// TIA Portal project "ND_PiPl" (V16)
// Lehrlingsprojekt

(* hardware
DEVICE "ET 200SP-Station_1"  ET 200SP-Station
   slot 0: "Baugruppenträger_0"  Rack  6ES5 710-8MAx1
   slot 1: "-20KF3"  CPU 1512SP F-1 PN  6ES7 512-1SK01-0AB0  V2.8
      slot 32768: "PROFINET-Schnittstelle_1"  X1
         slot 32771: "Port_3"  X1 P3
   slot 2: "-20KF5"  F-DI 8x24VDC HF  6ES7 136-6BA00-0CA0  V1.0
      slot 1: "-20KF5"  F-DI 8x24VDC HF
   slot 3: "-20KF6"  F-DQ 8x24VDC/0.5A PP HF  6ES7 136-6DC00-0CA0  V1.0
      slot 1: "-20KF6"  F-DQ 8x24VDC/0.5A PP HF
   slot 4: "-21KF1"  DI 16x24VDC ST  6ES7 131-6BH01-0BA0  V0.0
      slot 1: "-21KF1"  DI 16x24VDC ST
   slot 5: "-21KF4"  DQ 16x24VDC/0.5A ST  6ES7 132-6BH01-0BA0  V0.0
      slot 1: "-21KF4"  DQ 16x24VDC/0.5A ST
   slot 6: "-22KF1"  AI 2xU/I 2-,4-wire HS  6ES7 134-6HB00-0DA1  V2.0
      slot 1: "-22KF1"  AI 2xU/I 2-,4-wire HS
   slot 7: "-22KF3"  AQ 2xU ST  6ES7 135-6FB00-0BA1  V1.0
      slot 1: "-22KF3"  AQ 2xU ST
   slot 8: "Servermodul_1"  Server module  6ES7 193-6PA00-0AA0  V1.1
      slot 1: "Servermodul_1"  Server module
   slot 127: "BA 2xRJ45"  BA 2xRJ45  6ES7 193-6AR00-0AA0  V0.0
      slot 32769: "Port_1"  X1 P1  6ES7 193-6AR00-0AA0
      slot 32770: "Port_2"  X1 P2  6ES7 193-6AR00-0AA0
DEVICE "HMI_1"  KTP400 Comfort
   slot 0: "HMI_1"  KTP400 Comfort  6AV2 124-2DC01-0AX0  16.0.0.0
   slot 1: "HMI_RT_1"  KTP400 Comfort  6AV2 124-2DC01-0AX0  16.0.0.0
   slot 5: "HMI_1.IE_CP_1"  PROFINET Interface  16.0.0.0
      slot 1: "PROFINET Schnittstelle_1"  PROFINET Interface
         slot 1: "Port_1"  Port
   slot 7: "HMI_1.MPI/DP_CP_1"  MPI/DP Interface  16.0.0.0
*)

// ===== PLC "-20KF3"  CPU 1512SP F-1 PN =====
// protected blocks, not shown: "Main_Safety_RTG1", "Main_Safety_RTG1_DB"

VAR_GLOBAL   // PLC tag table "Standard-Variablentabelle"
   "FirstScan" AT %M1.0 : Bool;
   "DiagStatusUpdate" AT %M1.1 : Bool;
   "AlwaysTRUE" AT %M1.2 : Bool;
   "AlwaysFALSE" AT %M1.3 : Bool;
   "Clock_10Hz" AT %M50.0 : Bool;
   "Clock_5Hz" AT %M50.1 : Bool;
   "Clock_2.5Hz" AT %M50.2 : Bool;
   "Clock_2Hz" AT %M50.3 : Bool;
   "Clock_1.25Hz" AT %M50.4 : Bool;
   "Clock_1Hz" AT %M50.5 : Bool;
   "Clock_0.625Hz" AT %M50.6 : Bool;
   "Clock_0.5Hz" AT %M50.7 : Bool;
   "MaschineStart" AT %M900.0 : Bool;
   "Schritt_Förderband_Ein" AT %M900.1 : Bool;
   "Schritt_Vereinzelner_Ein" AT %M900.2 : Bool;
   "Vereinzler_Ein" AT %M1000.0 : Bool;
   "Schritt_Horizontalarm_Zurück" AT %M900.3 : Bool;
   "Schritt_Vakuum_Ein" AT %M900.4 : Bool;
   "VakuumSR" AT %M1000.1 : Bool;
   "Förderband_Merker" AT %M2000.0 : Bool;
   "Schritt_Vertikalarm_runter" AT %M900.5 : Bool;
   "Tag_2" AT %M1000.2 : Bool;
   "Schritt_Vertikalarm_oben" AT %M900.6 : Bool;
   "Schritt_Horizontalarm_vor" AT %M900.7 : Bool;
   "Schritt_VertikalarmDeckel_runter" AT %M901.0 : Bool;
   "Schritt_Vakuum_aus" AT %M901.1 : Bool;
   "Schritt_VertikalarmDeckelweg_oben" AT %M901.2 : Bool;
   "Schritt_HorizontalarmDeckel_zurück" AT %M901.3 : Bool;
   "Schritt_Vereinzler_aus" AT %M901.4 : Bool;
   "Schritt_Zurücksetzten_Anfang" AT %M901.5 : Bool;
   "Start_Impuls" AT %M200.1 : Bool;
   "Einmal_Start" AT %M2000.1 : Bool;
   "Stop_Speicher" AT %M2000.2 : Bool;
   "Deckler_Speicher" AT %M2000.3 : Bool;
   "Tag_1" AT %ED500 : Real;
   "Druck_Zu_Niedrig" AT %M2000.4 : Bool;
   "Druck_Zu_Hoch" AT %M2000.5 : Bool;
   "Prod_Count" AT %MW1200 : Int;
   "Prod_Count_Reset" AT %M300.0 : Bool;
END_VAR

VAR_GLOBAL   // PLC tag table "Systemflags"
   "System_Byte" AT %MB1 : Byte;   // Byte System
   "ME_PLC_First_Scan_Bit" AT %M1.0 : Bool;   // PLC First Scan Bit
   "ME_PLC_DiagStatusUpdate" AT %M1.1 : Bool;   // PLC Diagnostic Status Update
   "ME_PLC_TRUE" AT %M1.2 : Bool;   // PLC TRUE
   "ME_PLC_FALSE" AT %M1.3 : Bool;   // PLC FALSE
   "Clock_Byte" AT %MB50 : Byte;   // Byte PLC Clock
   "ME_PLC_Clock_0.1s" AT %M0.0 : Bool;   // PLC Clock 0.1s (10Hz )
   "ME_PLC_Clock_0.2s" AT %M0.1 : Bool;   // PLC Clock 0.2s (5Hz )
   "ME_PLC_Clock_0.4s" AT %M0.2 : Bool;   // PLC Clock 0.4s (2.5Hz )
   "ME_PLC_Clock_0.5s" AT %M0.3 : Bool;   // PLC Clock 0.5s (2Hz )
   "ME_PLC_Clock_0.8s" AT %M0.4 : Bool;   // PLC Clock 0.8s (1.25Hz )
   "ME_PLC_Clock_1.0s" AT %M0.5 : Bool;   // PLC Clock 1s (1Hz)
   "ME_PLC_Clock_1.6s" AT %M0.6 : Bool;   // PLC Clock 1.6s (0.625Hz )
   "ME_PLC_Clock_2.0s" AT %M0.7 : Bool;   // PLC Clock 2s (0.5Hz )
   "ME_PLC_FC_Test" AT %M2.0 : Bool;   // Testing Frequency Converters
   "ME_PLC_TRUE_to_do" AT %M2.2 : Bool;   // PLC TRUE to do
   "ME_PLC_FALSE_to_do" AT %M2.3 : Bool;   // PLC FALSE to do
   "ME_PLC_Led_Error" AT %M2.4 : Bool;   // PLC LED Error
   "ME_PLC_Led_Maint" AT %M2.5 : Bool;   // PLC LED Maintenance
   "ME_PLC_Startup_Rst" AT %M2.6 : Bool;   // PLC LED Startup Reset
   "ME_PLC_First_Scan_Bit_FC" AT %M2.1 : Bool;   // Call Frequency Converters
END_VAR

VAR_GLOBAL   // PLC tag table "IO-Pick&Placer"
   "CC_KF_FbEStop" AT %E0.0 : Bool;   // Rückmeldung Freigabe Not-Halt (81KF8)
   "PPTR_BG_InletPart" AT %E0.1 : Bool;   // Transportband Werkstück am Bandanfang (100BG1)
   "PPTR_BG_PartAtSep" AT %E0.2 : Bool;   // Transportband Werkstück am Vereinzeler (100BG2)
   "PPTR_BG_BackupPart" AT %E0.3 : Bool;   // Transportband Werkstück beim Bandende (100BG3)
   "PIPL_BG_CarrierRetracted" AT %E0.4 : Bool;   // Pick&Placer Schlitten eingefahren (120BG1)
   "PIPL_BG_CarrierExtended" AT %E0.5 : Bool;   // Pick&Placer Schlitten ausgefahren (120BG2)
   "PIPL_BG_SuctTop" AT %E0.6 : Bool;   // Pick&Placer Sauger oben (120BG3)
   "PIPL_BP_PartSuckedOn" AT %E0.7 : Bool;   // Pick&Placer Werkstück angesaugt (120PB4)
   "PIPL_Pa_SF_Reset" AT %E1.0 : Bool;   // Pick&Placer Bedienstelle Reset (160SF2)
   "PIPL_Pa_SF_Start" AT %E1.1 : Bool;   // Pick&Placer Bedienstelle Start (160SF3)
   "PIPL_Pa_SF_Stop" AT %E1.2 : Bool;   // Pick&Placer Bedienstelle Stop (160SF4)
   "PIPL_Pa_SF_ManAuto" AT %E1.3 : Bool;   // Pick&Placer Bedienstelle Manual - Auto (160SF5)
   "CC_Spare_I1.4" AT %E1.4 : Bool;   // Spare
   "CC_Spare_I1.5" AT %E1.5 : Bool;   // Spare
   "CC_Spare_I1.6" AT %E1.6 : Bool;   // Spare
   "CC_Spare_I1.7" AT %E1.7 : Bool;   // Spare
   "PPTR_MB_SeparatorExtend" AT %A0.0 : Bool;   // Transportband Vereinzeler ausfahren (105MB8)
   "PIPL_SC_Green" AT %A0.1 : Bool;   // Pick&Placer Turmleuchte grün (130PF1)
   "PIPL_SC_Yellow" AT %A0.2 : Bool;   // Pick&Placer Turmleuchte gelb (130PF1)
   "PIPL_SC_Red" AT %A0.3 : Bool;   // Pick&Placer Turmleuchte rot (130PF1)
   "PIPL_MB_CarrierExtend" AT %A0.4 : Bool;   // Pick&Placer Schlitten ausfahren (125MB1)
   "PIPL_MB_CarrierRetract" AT %A0.5 : Bool;   // Pick&Placer Schlitten einfahren (125MB2)
   "PIPL_MB_SuctDown" AT %A0.6 : Bool;   // Pick&Placer Sauger nach unten (125MB3)
   "PIPL_MB_VacuumOn" AT %A0.7 : Bool;   // Pick&Placer Vakuum ein (125MB4)
   "PIPL_Pa_PF_ControlCircuit" AT %A1.0 : Bool;   // Pick&Placer Bedienstelle LED Steuerspannung Ein (Reset) (160SF2)
   "PIPL_Pa_PF_Error" AT %A1.1 : Bool;   // Pick&Placer Bedienstelle LED Fehler (160PF2)
   "PIPL_Pa_PF_Start" AT %A1.2 : Bool;   // Pick&Placer Bedienstelle LED Start (160SF3)
   "CC_Spare_O1.3" AT %A1.3 : Bool;   // Spare
   "CC_Spare_O1.4" AT %A1.4 : Bool;   // Spare
   "CC_Spare_O1.5" AT %A1.5 : Bool;   // Spare
   "CC_Spare_O1.6" AT %A1.6 : Bool;   // Spare
   "CC_Spare_O1.7" AT %A1.7 : Bool;   // Spare
   "Druck_Tester" AT %EW272 : Int;   // Druck Tester
   "CC_Spare_IW274" AT %EW274 : Word;   // Spare
   "PPTR_TF_DriveSpeed" AT %AW272 : Word;   // Transportband Bandmotor Geschwindigkeit Option (105TF1)
   "CC_Spare_OW274" AT %AW274 : Word;   // Spare
   "Druck_Zwischenwert" AT %MD276 : Real;
   "Druck_Wert1" AT %MD280 : Real;
   "Druck_Wert2" AT %MW284 : Int;
   "Druck_Wert_Final" AT %MD286 : Real;
END_VAR

VAR_GLOBAL   // PLC tag table "IO-Pick&Placer-Safety"
   "PIPL_Pa_EStopCh1" AT %E1000.0 : Bool;   // Pick&Placer Bedienstelle Not-Halt Channel 1 (160SF1)
   "CC_Spare_I1000.1" AT %E1000.1 : Bool;   // Spare
   "CC_Spare_I1000.2" AT %E1000.2 : Bool;   // Spare
   "CC_Spare_I1000.3" AT %E1000.3 : Bool;   // Spare
   "PIPL_Pa_EStopCh2" AT %E1000.4 : Bool;   // Pick&Placer Bedienstelle Not-Halt Channel 2 (160SF1)
   "CC_Spare_I1000.5" AT %E1000.5 : Bool;   // Spare
   "CC_Spare_I1000.6" AT %E1000.6 : Bool;   // Spare
   "CC_Spare_I1000.7" AT %E1000.7 : Bool;   // Spare
   "CC_KF_EStopCh1" AT %A1050.0 : Bool;   // Freigabe Not-Halt Channel 1 (81KF7)
   "CC_KF_EStopCh2" AT %A1050.1 : Bool;   // Freigabe Not-Halt Channel 2 (81KF8)
   "PPTR_TF_DriveForward" AT %A1050.2 : Bool;   // Transportband Bandmotor Vorwärts (105TF1)
   "PPTR_TF_DriveReverse" AT %A1050.3 : Bool;   // Transportband Bandmotor Rückwärts (105TF1)
   "CC_Spare_O1050.4" AT %A1050.4 : Bool;   // Spare
   "CC_Spare_O1050.5" AT %A1050.5 : Bool;   // Spare
   "CC_Spare_O1050.6" AT %A1050.6 : Bool;   // Spare
   "CC_Spare_O1050.7" AT %A1050.7 : Bool;   // Spare
END_VAR

DATA_BLOCK "HMI_Meldungen"   // DB120
{ S7_Optimized_Access := 'FALSE' }
VERSION : 0.1
   VAR
      Fehler : Struct
         "Not-Aus" : Bool;   // NOT-Aus Aktiv
         "Not-Aus_Quit" : Bool;   // NOT-Aus Quitieren
         "2" : Bool;
         "3" : Bool;
         "4" : Bool;
         "5" : Bool;
         "6" : Bool;
         "7" : Bool;
         "8" : Bool;
         "9" : Bool;
         "10" : Bool;
         "11" : Bool;
         "12" : Bool;
         "13" : Bool;
         "14" : Bool;
         "15" : Bool;
      END_STRUCT;
      Meldungen : Struct
         "0" : Bool;
         "1" : Bool;
         "2" : Bool;
         "3" : Bool;
         "4" : Bool;
         "5" : Bool;
         "6" : Bool;
         "7" : Bool;
         "8" : Bool;
         "9" : Bool;
         "10" : Bool;
         "11" : Bool;
         "12" : Bool;
         "13" : Bool;
         "14" : Bool;
         "15" : Bool;
      END_STRUCT;
      Warnungen : Struct
         Druck_zu_niedrig : Bool;   // Druck zu niedrig
         Druck_zu_hoch : Bool;   // Druck zu hoch
         Keine_Deckel : Bool;   // Keine Deckel vorhanden
         Rückstau : Bool;   // Rückstau am Bandende
         "4" : Bool;
         "5" : Bool;
         "6" : Bool;
         "7" : Bool;
         "8" : Bool;
         "9" : Bool;
         "10" : Bool;
         "11" : Bool;
         "12" : Bool;
         "13" : Bool;
         "14" : Bool;
         "15" : Bool;
      END_STRUCT;
   END_VAR
BEGIN
END_DATA_BLOCK

// folder: System blocks/Program resources

DATA_BLOCK "IEC_Timer_0_DB"   // DB3
{ S7_Optimized_Access := 'TRUE' }
AUTHOR : Simatic
FAMILY : IEC
NAME : IEC_TMR
VERSION : 1.0
// stored: InstanceOfName IEC_TIMER
"IEC_TIMER"
BEGIN
END_DATA_BLOCK

DATA_BLOCK "Vakuum_Timer_Ausschalten"   // DB5
{ S7_Optimized_Access := 'TRUE' }
AUTHOR : Simatic
FAMILY : IEC
NAME : IEC_TMR
VERSION : 1.0
// stored: InstanceOfName IEC_TIMER
"IEC_TIMER"
BEGIN
END_DATA_BLOCK

DATA_BLOCK "Timer_Rückstau"   // DB6
{ S7_Optimized_Access := 'TRUE' }
AUTHOR : Simatic
FAMILY : IEC
NAME : IEC_TMR
VERSION : 1.0
// stored: InstanceOfName IEC_TIMER
"IEC_TIMER"
BEGIN
END_DATA_BLOCK

DATA_BLOCK "Timer_Clean_Reset"   // DB7
{ S7_Optimized_Access := 'TRUE' }
AUTHOR : Simatic
FAMILY : IEC
NAME : IEC_TMR
VERSION : 1.0
// stored: InstanceOfName IEC_TIMER
"IEC_TIMER"
BEGIN
END_DATA_BLOCK

DATA_BLOCK "IEC_Counter_0_DB"   // DB8
{ S7_Optimized_Access := 'TRUE' }
AUTHOR : Simatic
FAMILY : IEC
NAME : CNTR
VERSION : 1.0
// stored: InstanceOfName IEC_COUNTER
"IEC_COUNTER"
BEGIN
END_DATA_BLOCK

// folder: (top level)

FUNCTION "Ausgänge" : Void   // FC1, FBD
{ S7_Optimized_Access := 'TRUE' }
VERSION : 0.1
BEGIN

REGION Network 1: Vereinzler
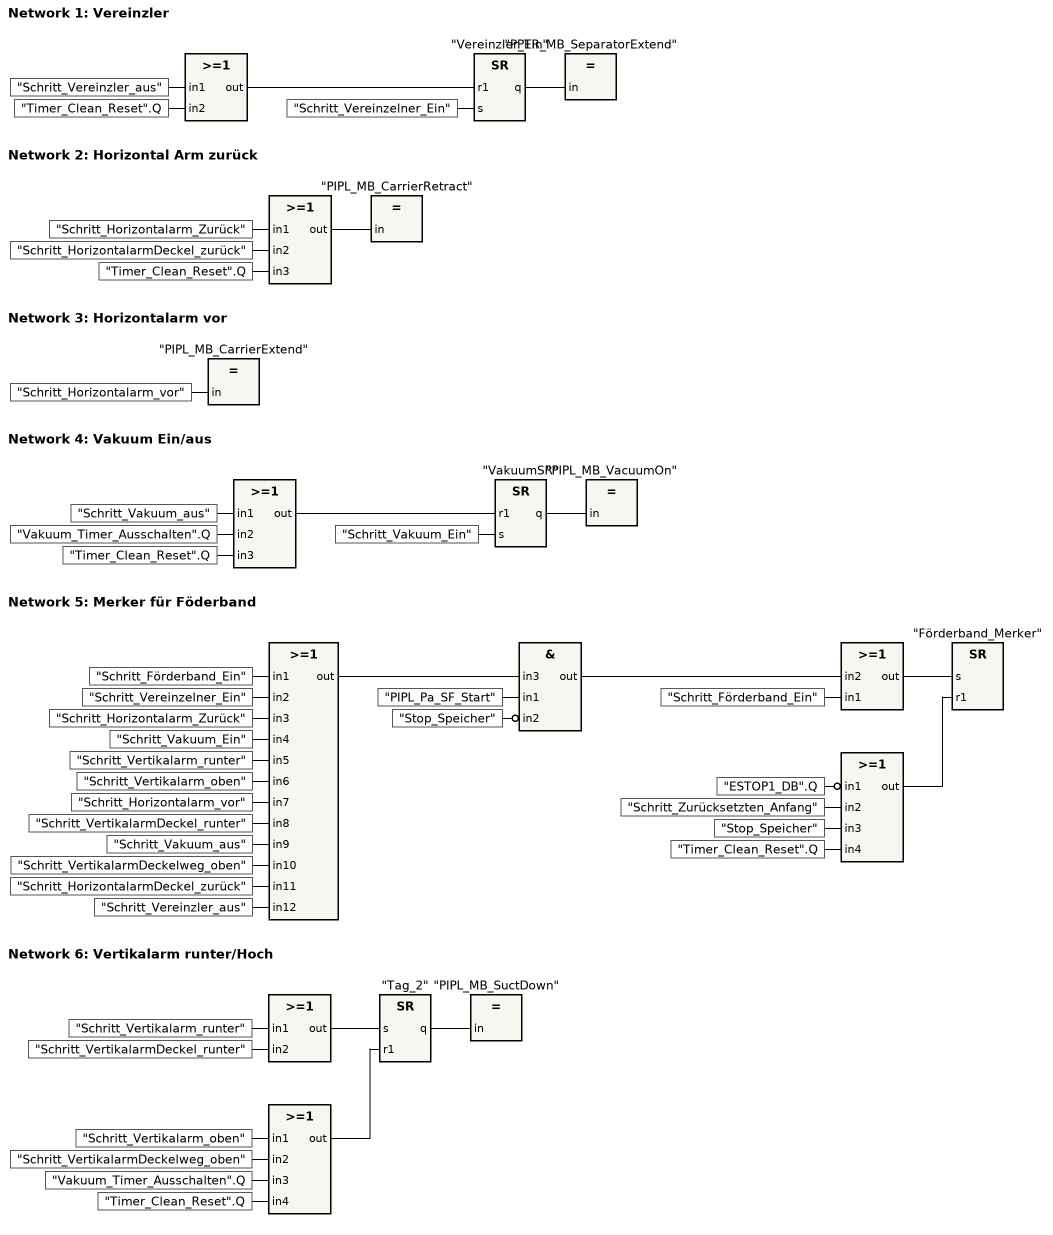
   IF "Schritt_Vereinzelner_Ein" THEN
       "Vereinzler_Ein" := TRUE;   // SR flip-flop
   END_IF;
   IF "Schritt_Vereinzler_aus" OR "Timer_Clean_Reset".Q THEN "Vereinzler_Ein" := FALSE; END_IF;
   "PPTR_MB_SeparatorExtend" := "Vereinzler_Ein";
END_REGION

REGION Network 2: Horizontal Arm zurück
   "PIPL_MB_CarrierRetract" := "Schritt_Horizontalarm_Zurück" OR "Schritt_HorizontalarmDeckel_zurück" OR "Timer_Clean_Reset".Q;
END_REGION

REGION Network 3: Horizontalarm vor
   "PIPL_MB_CarrierExtend" := "Schritt_Horizontalarm_vor";
END_REGION

REGION Network 4: Vakuum Ein/aus
   IF "Schritt_Vakuum_Ein" THEN
       "VakuumSR" := TRUE;   // SR flip-flop
   END_IF;
   IF "Schritt_Vakuum_aus" OR "Vakuum_Timer_Ausschalten".Q OR "Timer_Clean_Reset".Q THEN
       "VakuumSR" := FALSE;
   END_IF;
   "PIPL_MB_VacuumOn" := "VakuumSR";
END_REGION

REGION Network 5: Merker für Föderband
   IF (("Schritt_Förderband_Ein" OR "Schritt_Vereinzelner_Ein" OR "Schritt_Horizontalarm_Zurück" OR "Schritt_Vakuum_Ein" OR "Schritt_Vertikalarm_runter" OR "Schritt_Vertikalarm_oben" OR "Schritt_Horizontalarm_vor" OR "Schritt_VertikalarmDeckel_runter" OR "Schritt_Vakuum_aus" OR "Schritt_VertikalarmDeckelweg_oben" OR "Schritt_HorizontalarmDeckel_zurück" OR "Schritt_Vereinzler_aus") AND "PIPL_Pa_SF_Start" AND NOT "Stop_Speicher") OR "Schritt_Förderband_Ein" THEN
       "Förderband_Merker" := TRUE;   // SR flip-flop
   END_IF;
   IF NOT "ESTOP1_DB".Q OR "Schritt_Zurücksetzten_Anfang" OR "Stop_Speicher" OR "Timer_Clean_Reset".Q THEN
       "Förderband_Merker" := FALSE;
   END_IF;
END_REGION

REGION Network 6: Vertikalarm runter/Hoch
   IF "Schritt_Vertikalarm_runter" OR "Schritt_VertikalarmDeckel_runter" THEN
       "Tag_2" := TRUE;   // SR flip-flop
   END_IF;
   IF "Schritt_Vertikalarm_oben" OR "Schritt_VertikalarmDeckelweg_oben" OR "Vakuum_Timer_Ausschalten".Q OR "Timer_Clean_Reset".Q THEN
       "Tag_2" := FALSE;
   END_IF;
   "PIPL_MB_SuctDown" := "Tag_2";
END_REGION
END_FUNCTION

FUNCTION "Pick&Place_Auto" : Void   // FC2, FBD
{ S7_Optimized_Access := 'TRUE' }
VERSION : 0.1
BEGIN

REGION Network 1: Eischalten der Maschine
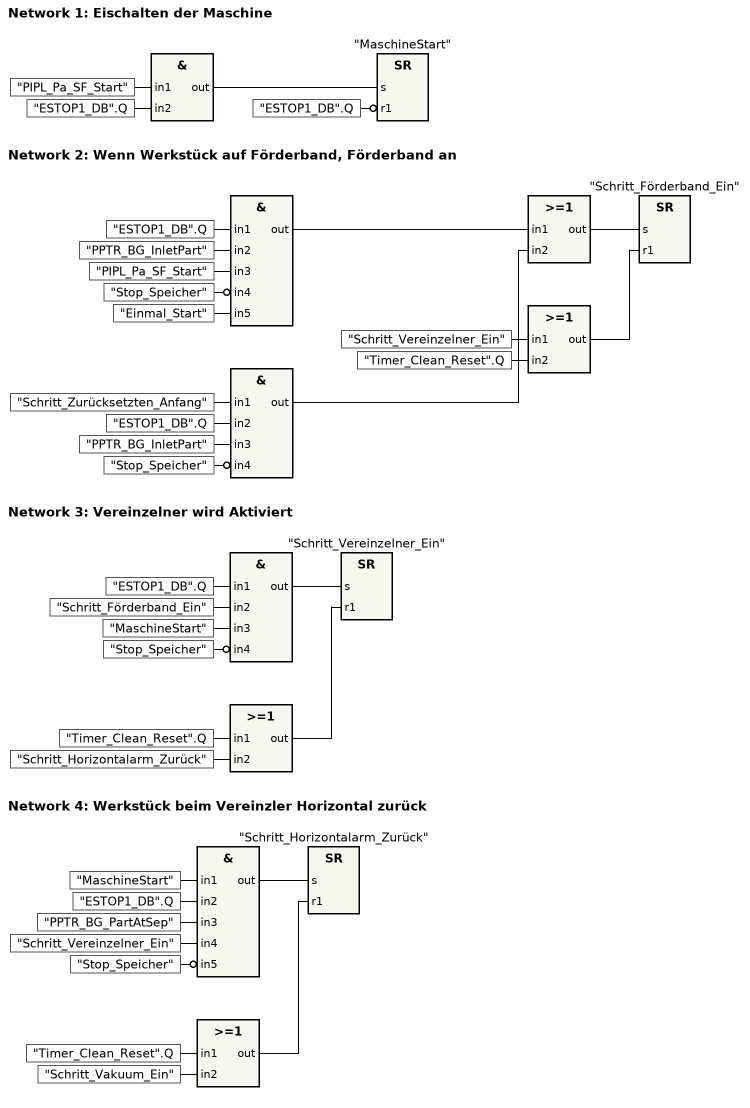
   IF "PIPL_Pa_SF_Start" AND "ESTOP1_DB".Q THEN
       "MaschineStart" := TRUE;   // SR flip-flop
   END_IF;
   IF NOT "ESTOP1_DB".Q THEN "MaschineStart" := FALSE; END_IF;
END_REGION

REGION Network 2: Wenn Werkstück auf Förderband, Förderband an
   IF ("ESTOP1_DB".Q AND "PPTR_BG_InletPart" AND "PIPL_Pa_SF_Start" AND NOT "Stop_Speicher" AND "Einmal_Start") OR ("Schritt_Zurücksetzten_Anfang" AND "ESTOP1_DB".Q AND "PPTR_BG_InletPart" AND NOT "Stop_Speicher") THEN
       "Schritt_Förderband_Ein" := TRUE;   // SR flip-flop
   END_IF;
   IF "Schritt_Vereinzelner_Ein" OR "Timer_Clean_Reset".Q THEN "Schritt_Förderband_Ein" := FALSE; END_IF;
END_REGION

REGION Network 3: Vereinzelner wird Aktiviert
   IF "ESTOP1_DB".Q AND "Schritt_Förderband_Ein" AND "MaschineStart" AND NOT "Stop_Speicher" THEN
       "Schritt_Vereinzelner_Ein" := TRUE;   // SR flip-flop
   END_IF;
   IF "Timer_Clean_Reset".Q OR "Schritt_Horizontalarm_Zurück" THEN
       "Schritt_Vereinzelner_Ein" := FALSE;
   END_IF;
END_REGION

REGION Network 4: Werkstück beim Vereinzler Horizontal zurück
   IF "MaschineStart" AND "ESTOP1_DB".Q AND "PPTR_BG_PartAtSep" AND "Schritt_Vereinzelner_Ein" AND NOT "Stop_Speicher" THEN
       "Schritt_Horizontalarm_Zurück" := TRUE;   // SR flip-flop
   END_IF;
   IF "Timer_Clean_Reset".Q OR "Schritt_Vakuum_Ein" THEN "Schritt_Horizontalarm_Zurück" := FALSE; END_IF;
END_REGION

REGION Network 5: Wenn Horizontalarm zurück, Vakuum ein
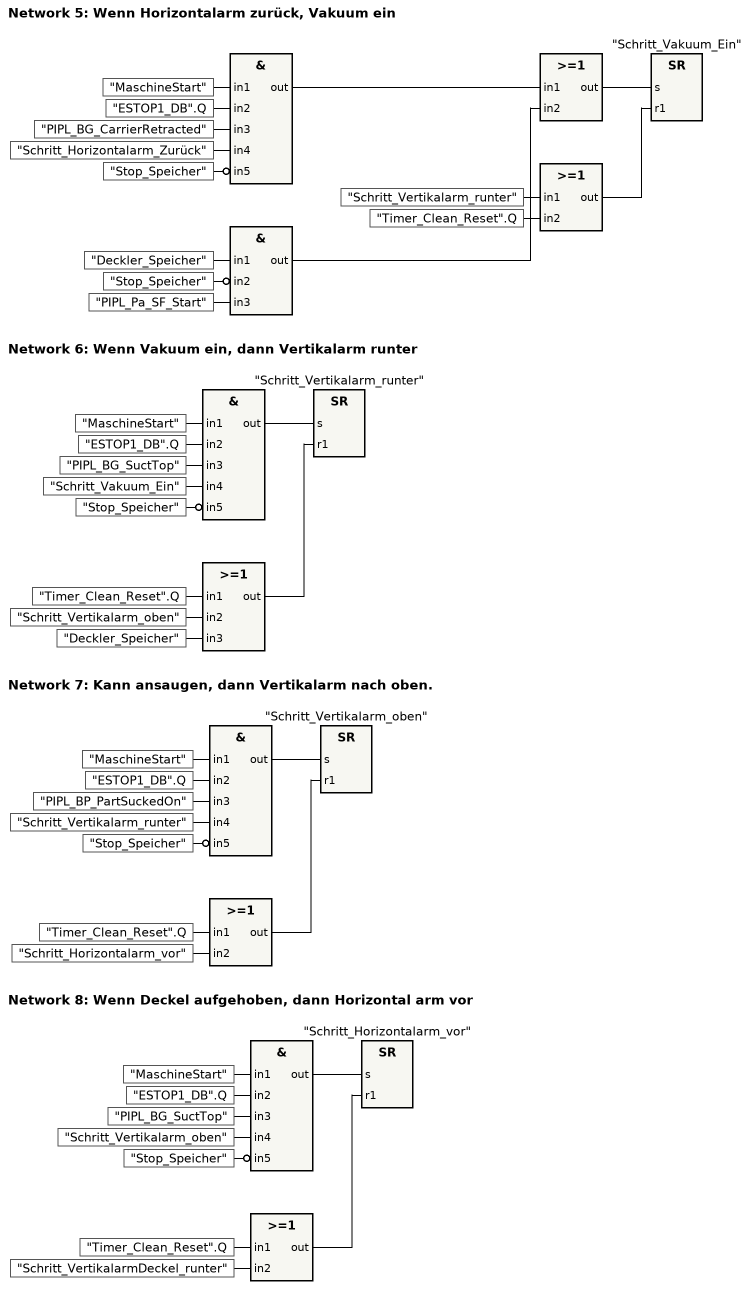
   IF ("MaschineStart" AND "ESTOP1_DB".Q AND "PIPL_BG_CarrierRetracted" AND "Schritt_Horizontalarm_Zurück" AND NOT "Stop_Speicher") OR ("Deckler_Speicher" AND NOT "Stop_Speicher" AND "PIPL_Pa_SF_Start") THEN
       "Schritt_Vakuum_Ein" := TRUE;   // SR flip-flop
   END_IF;
   IF "Schritt_Vertikalarm_runter" OR "Timer_Clean_Reset".Q THEN "Schritt_Vakuum_Ein" := FALSE; END_IF;
END_REGION

REGION Network 6: Wenn Vakuum ein, dann Vertikalarm runter
   IF "MaschineStart" AND "ESTOP1_DB".Q AND "PIPL_BG_SuctTop" AND "Schritt_Vakuum_Ein" AND NOT "Stop_Speicher" THEN
       "Schritt_Vertikalarm_runter" := TRUE;   // SR flip-flop
   END_IF;
   IF "Timer_Clean_Reset".Q OR "Schritt_Vertikalarm_oben" OR "Deckler_Speicher" THEN
       "Schritt_Vertikalarm_runter" := FALSE;
   END_IF;
END_REGION

REGION Network 7: Kann ansaugen, dann Vertikalarm nach oben.
   IF "MaschineStart" AND "ESTOP1_DB".Q AND "PIPL_BP_PartSuckedOn" AND "Schritt_Vertikalarm_runter" AND NOT "Stop_Speicher" THEN
       "Schritt_Vertikalarm_oben" := TRUE;   // SR flip-flop
   END_IF;
   IF "Timer_Clean_Reset".Q OR "Schritt_Horizontalarm_vor" THEN "Schritt_Vertikalarm_oben" := FALSE; END_IF;
END_REGION

REGION Network 8: Wenn Deckel aufgehoben, dann Horizontal arm vor
   IF "MaschineStart" AND "ESTOP1_DB".Q AND "PIPL_BG_SuctTop" AND "Schritt_Vertikalarm_oben" AND NOT "Stop_Speicher" THEN
       "Schritt_Horizontalarm_vor" := TRUE;   // SR flip-flop
   END_IF;
   IF "Timer_Clean_Reset".Q OR "Schritt_VertikalarmDeckel_runter" THEN
       "Schritt_Horizontalarm_vor" := FALSE;
   END_IF;
END_REGION

REGION Network 9: Wenn Horizontalarm vor mit Deckel, dann Vertickalarm runter
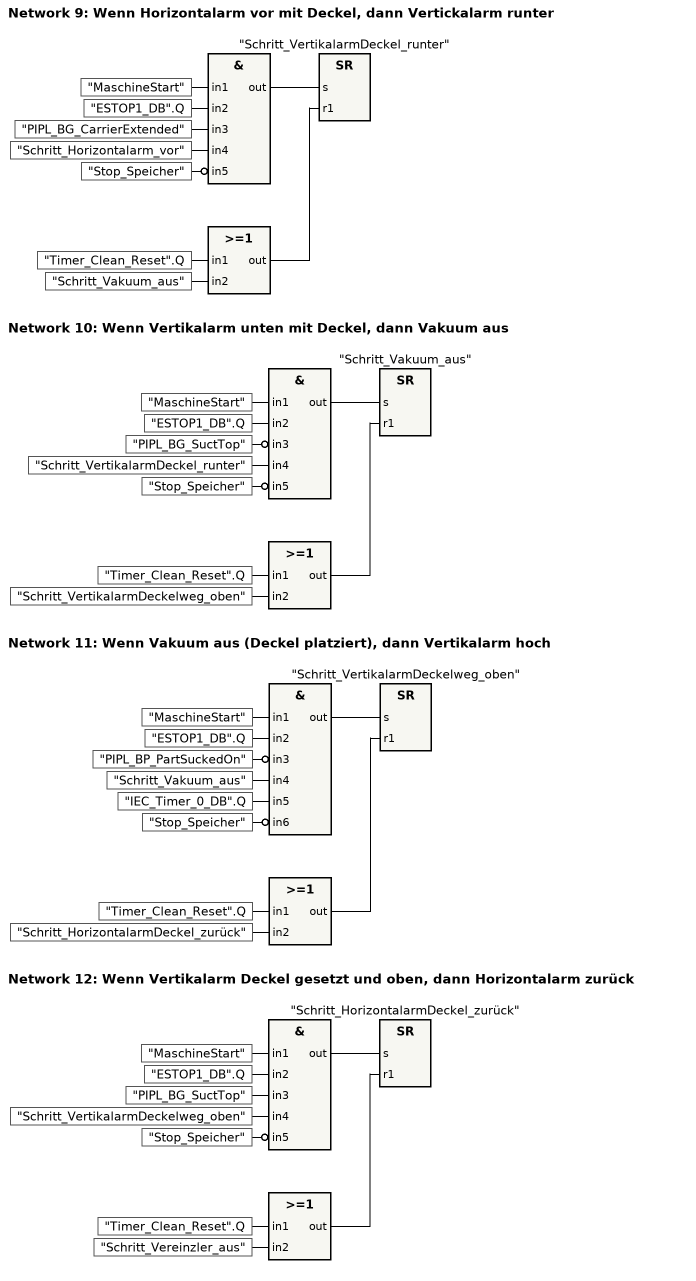
   IF "MaschineStart" AND "ESTOP1_DB".Q AND "PIPL_BG_CarrierExtended" AND "Schritt_Horizontalarm_vor" AND NOT "Stop_Speicher" THEN
       "Schritt_VertikalarmDeckel_runter" := TRUE;   // SR flip-flop
   END_IF;
   IF "Timer_Clean_Reset".Q OR "Schritt_Vakuum_aus" THEN "Schritt_VertikalarmDeckel_runter" := FALSE; END_IF;
END_REGION

REGION Network 10: Wenn Vertikalarm unten mit Deckel, dann Vakuum aus
   IF "MaschineStart" AND "ESTOP1_DB".Q AND NOT "PIPL_BG_SuctTop" AND "Schritt_VertikalarmDeckel_runter" AND NOT "Stop_Speicher" THEN
       "Schritt_Vakuum_aus" := TRUE;   // SR flip-flop
   END_IF;
   IF "Timer_Clean_Reset".Q OR "Schritt_VertikalarmDeckelweg_oben" THEN
       "Schritt_Vakuum_aus" := FALSE;
   END_IF;
END_REGION

REGION Network 11: Wenn Vakuum aus (Deckel platziert), dann Vertikalarm hoch
   IF "MaschineStart" AND "ESTOP1_DB".Q AND NOT "PIPL_BP_PartSuckedOn" AND "Schritt_Vakuum_aus" AND "IEC_Timer_0_DB".Q AND NOT "Stop_Speicher" THEN
       "Schritt_VertikalarmDeckelweg_oben" := TRUE;   // SR flip-flop
   END_IF;
   IF "Timer_Clean_Reset".Q OR "Schritt_HorizontalarmDeckel_zurück" THEN
       "Schritt_VertikalarmDeckelweg_oben" := FALSE;
   END_IF;
END_REGION

REGION Network 12: Wenn Vertikalarm Deckel gesetzt und oben, dann Horizontalarm zurück
   IF "MaschineStart" AND "ESTOP1_DB".Q AND "PIPL_BG_SuctTop" AND "Schritt_VertikalarmDeckelweg_oben" AND NOT "Stop_Speicher" THEN
       "Schritt_HorizontalarmDeckel_zurück" := TRUE;   // SR flip-flop
   END_IF;
   IF "Timer_Clean_Reset".Q OR "Schritt_Vereinzler_aus" THEN
       "Schritt_HorizontalarmDeckel_zurück" := FALSE;
   END_IF;
END_REGION

REGION Network 13: Wenn Horizontalarm zurück (Deckel platziert), dann Vereinzler aus
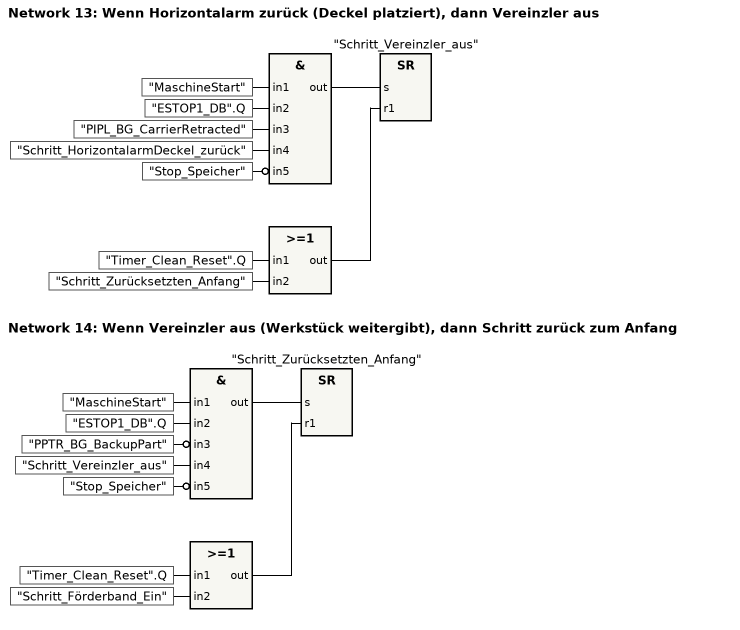
   IF "MaschineStart" AND "ESTOP1_DB".Q AND "PIPL_BG_CarrierRetracted" AND "Schritt_HorizontalarmDeckel_zurück" AND NOT "Stop_Speicher" THEN
       "Schritt_Vereinzler_aus" := TRUE;   // SR flip-flop
   END_IF;
   IF "Timer_Clean_Reset".Q OR "Schritt_Zurücksetzten_Anfang" THEN "Schritt_Vereinzler_aus" := FALSE; END_IF;
END_REGION

REGION Network 14: Wenn Vereinzler aus (Werkstück weitergibt), dann Schritt zurück zum Anfang
   IF "MaschineStart" AND "ESTOP1_DB".Q AND NOT "PPTR_BG_BackupPart" AND "Schritt_Vereinzler_aus" AND NOT "Stop_Speicher" THEN
       "Schritt_Zurücksetzten_Anfang" := TRUE;   // SR flip-flop
   END_IF;
   IF "Timer_Clean_Reset".Q OR "Schritt_Förderband_Ein" THEN "Schritt_Zurücksetzten_Anfang" := FALSE; END_IF;
END_REGION
END_FUNCTION

FUNCTION "SonderBlöcke" : Void   // FC3, FBD
{ S7_Optimized_Access := 'TRUE' }
VERSION : 0.1
BEGIN

REGION Network 1: Delay für Deckel setzen
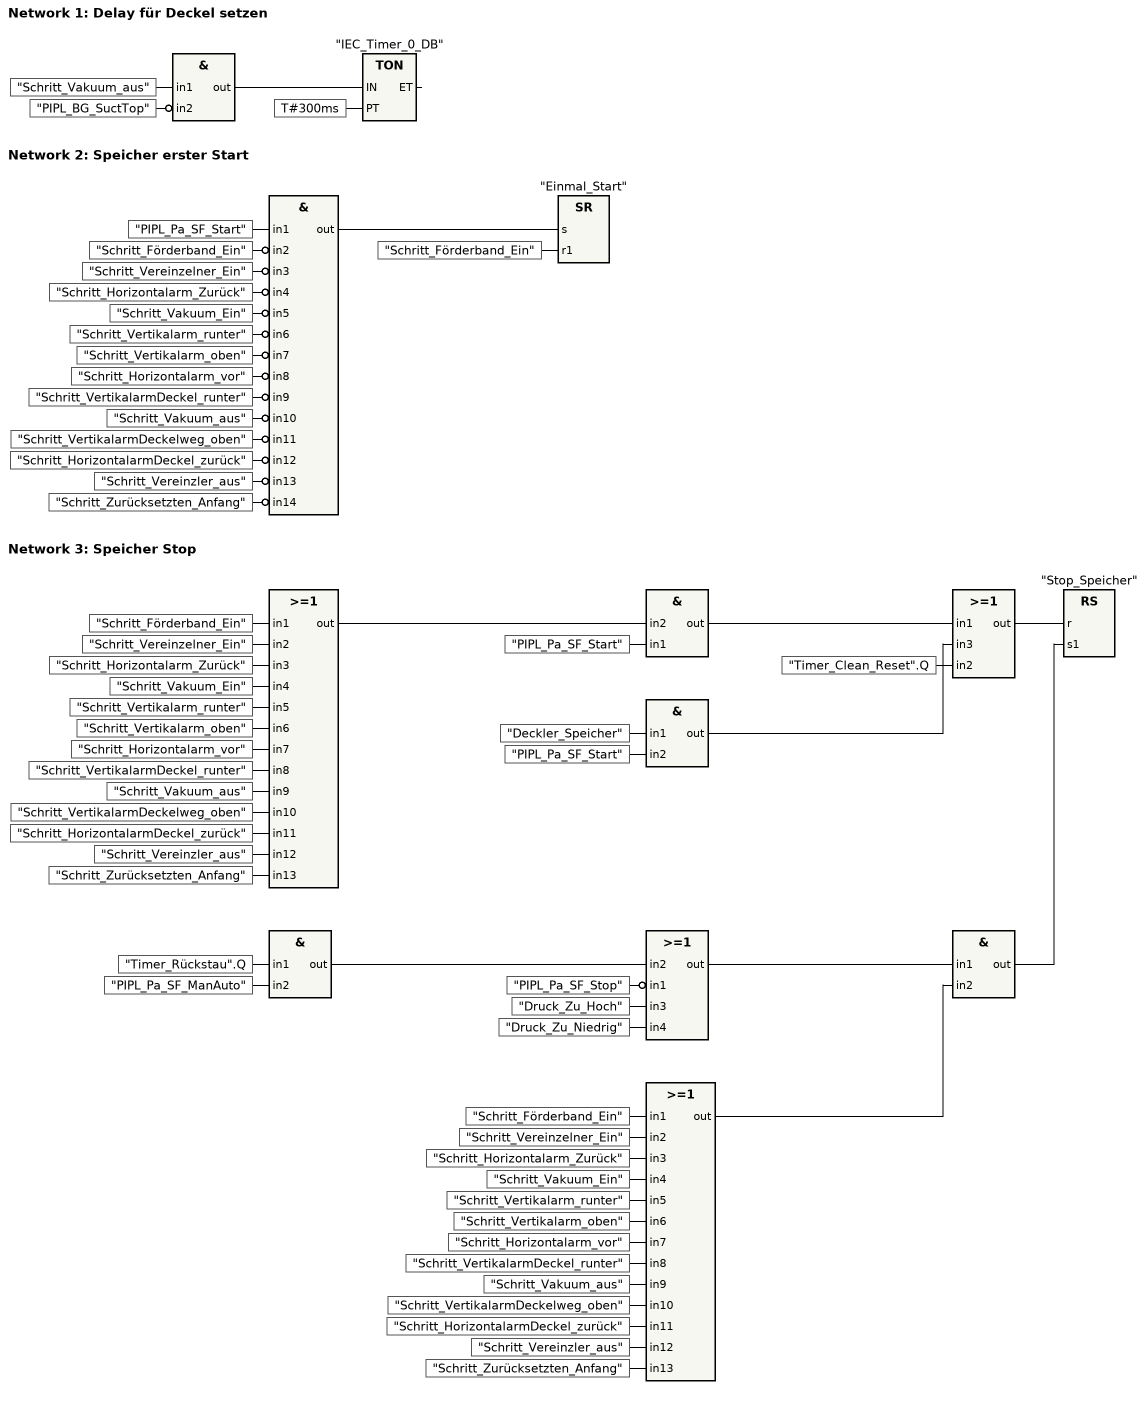
   "IEC_Timer_0_DB".TON(IN := "Schritt_Vakuum_aus" AND NOT "PIPL_BG_SuctTop", PT := T#300ms);
END_REGION

REGION Network 2: Speicher erster Start
   IF "PIPL_Pa_SF_Start" AND NOT "Schritt_Förderband_Ein" AND NOT "Schritt_Vereinzelner_Ein" AND NOT "Schritt_Horizontalarm_Zurück" AND NOT "Schritt_Vakuum_Ein" AND NOT "Schritt_Vertikalarm_runter" AND NOT "Schritt_Vertikalarm_oben" AND NOT "Schritt_Horizontalarm_vor" AND NOT "Schritt_VertikalarmDeckel_runter" AND NOT "Schritt_Vakuum_aus" AND NOT "Schritt_VertikalarmDeckelweg_oben" AND NOT "Schritt_HorizontalarmDeckel_zurück" AND NOT "Schritt_Vereinzler_aus" AND NOT "Schritt_Zurücksetzten_Anfang" THEN
       "Einmal_Start" := TRUE;   // SR flip-flop
   END_IF;
   IF "Schritt_Förderband_Ein" THEN "Einmal_Start" := FALSE; END_IF;
END_REGION
